// TIA Portal project "1905391_001_000" (V16)

(* hardware
DEVICE "S7-1200 station_1"  S7-1200 Station
   slot 0: "Rack_0"  S7-1200 Rack  Rack  V1.0
   slot 1: "PLC_1"  CPU 1212C DC/DC/Rly  6ES7 212-1HE40-0XB0  V4.4
DEVICE "HMI_1"  TP900 Comfort
   slot 0: "HMI_1"  TP900 Comfort  6AV2 124-0JC01-0AX0  16.0.0.0
   slot 1: "HMI_RT_1"  TP900 Comfort  6AV2 124-0JC01-0AX0  16.0.0.0
   slot 5: "HMI_1.IE_CP_1"  PROFINET Interface  16.0.0.0
      slot 1: "PROFINET Interface_1"  PROFINET Interface
         slot 1: "Port_1"  Port
         slot 2: "Port_2"  Port
   slot 7: "HMI_1.MPI/DP_CP_1"  MPI/DP Interface  16.0.0.0
*)

// ===== PLC "PLC_1"  CPU 1212C DC/DC/Rly =====

VAR_GLOBAL   // PLC tag table "Default tag table"
   "System_Byte" AT %MB1 : Byte;
   "FirstScan" AT %M1.0 : Bool;
   "DiagStatusUpdate" AT %M1.1 : Bool;
   "AlwaysTRUE" AT %M1.2 : Bool;
   "AlwaysFALSE" AT %M1.3 : Bool;
   "Clock_Byte" AT %MB0 : Byte;
   "Clock_10Hz" AT %M0.0 : Bool;
   "Clock_5Hz" AT %M0.1 : Bool;
   "Clock_2.5Hz" AT %M0.2 : Bool;
   "Clock_2Hz" AT %M0.3 : Bool;
   "Clock_1.25Hz" AT %M0.4 : Bool;
   "Clock_1Hz" AT %M0.5 : Bool;
   "Clock_0.625Hz" AT %M0.6 : Bool;
   "Clock_0.5Hz" AT %M0.7 : Bool;
END_VAR

VAR_GLOBAL CONSTANT   // PLC tag table "Default tag table"
   "STRING_LENGTH" : Int := 20;
   "ADP_PARAMETER_LENGTH" : Int := 5;
   "NULL_TOKEN" : Int := -1;
   "BUSY_INDICATOR_OFF" : String := '200;200;200';
   "BUSY_INDICATOR_ON" : String := '250;250;150';
   "ERROR_INDICATOR_OFF" : String := '200;200;200';
   "ERROR_INDICATOR_ON" : String := '250;150;150';
   "STATUS_CODE_OFF" : String := '200;200;200';
   "OPERATION_LABEL_OFF" : String := '200;200;200';
   "CONNECTION_STATUS_HEADER" : String := '200;200;200';
   "STATUS_CODE_PROBLEM" : String := '250;150;150';
   "STATUS_CODE_GOOD" : String := '150;250;150';
END_VAR

VAR_GLOBAL CONSTANT   // PLC tag table "Colors"
   "LABEL_COLOR" : String := '200_200_200';
   "DESELECTED_INPUT_COLOR" : String := '250_250_250';
   "SELECTED_INPUT_COLOR" : String := '150,250,150';
   "BORDER_COLOR" : String := '200_200_200';
   "DIVIDER_COLOR" : String := '50_75_100';
   "THIS_SCREEN_COLOR" : String := '150;150;150';
   "OTHER_SCREEN_COLOR" : String := '100,100,100';
   "ACTUATE" : String := '150_250_150';
   "BACKGROUND_COLOR" : String := '150,150,200';
   "DONE_INDICATOR_OFF" : String := '200;200;200';
   "DONE_INDICATOR_ON" : String := '150;250;150';
   "OPERATION_OFF" : String := '200;200;200';
END_VAR

VAR_GLOBAL CONSTANT   // PLC tag table "Screen_Numbers"
   "WIRE_SCREEN_NUMBER" : Int := 1;
   "MATERIAL_SCREEN_NUMBER" : Int := 2;
   "CONNECTION_CONTROLS_SCREEN_NUMBER" : Int := 3;
   "CONNECTION_STATUS_DETAILS_SCREEN_NUMBER" : Int := 4;
   "CONNECTION_PARAMETERS_SCREEN_NUMBER" : Int := 5;
END_VAR

VAR_GLOBAL CONSTANT   // PLC tag table "Parameter_Entry_Modes"
   "MATERIAL" : String := 'MATERIAL';
   "WIRE" : String := 'WIRE';
END_VAR

VAR_GLOBAL CONSTANT   // PLC tag table "Connection_Statuses"
   "IDLE" : Word := 16#7000;
   "SUCCESS" : Word := 0;
END_VAR

VAR_GLOBAL CONSTANT   // PLC tag table "Send_Modes"
   "MANUAL" : String := 'MANUAL';
   "AUTOMATIC" : String := 'AUTOMATIC';
END_VAR

VAR_GLOBAL CONSTANT   // PLC tag table "Connection_Modes"
   "DISCONNECT_SELECTOR" : DInt := 1;
   "CONNECT_SELECTOR" : DInt := 2;
   "SEND_SELECTOR" : DInt := 3;
   "MATERIAL_DISCONNECT" : DInt := 1;
   "MATERIAL_CONNECT" : DInt := 2;
   "MATERIAL_SEND" : DInt := 3;
   "WIRE_DISCONNECT" : DInt := 4;
   "WIRE_CONNECT" : DInt := 5;
   "WIRE_SEND" : DInt := 6;
END_VAR

TYPE "Divider.UDT"
   STRUCT
      background_animate : DInt;
      background_visible : Bool;
      line_animate : DInt;
      line_visible : Bool;
   END_STRUCT;
END_TYPE

TYPE "Row_Data.UDT"
   STRUCT
      background_animate : DInt;
      background_visible : Bool;
      cell_0_animate : DInt;
      cell_0_visible : Bool;
      cell_1_active : Bool;
      cell_1_animate : DInt;
      cell_1_enable : Bool;
      cell_1_input_finished : Bool;
      cell_1_value : String[50];
      cell_1_visible : Bool;
   END_STRUCT;
END_TYPE

TYPE "HMI_Interface.UDT"
   STRUCT
      connection_parameters : "Connection_Paramters_HMI.UDT";
      connection_status_details : "Connection_Detail.HMI.UDT";
      connection_controls : "Connection_Status.HMI.UDT";
      materials : "Materials.HMI.UDT";
      meta : "HMI_Meta.UDT";
      navigation : "Navigation.HMI.UDT";
      wires : "Wire.HMI.UDT";
   END_STRUCT;
END_TYPE

TYPE "Navigation.HMI.UDT"
   STRUCT
      background_animate : DInt;
      background_visible : Bool;
      bottom_line_animate : DInt;
      bottom_line_visible : Bool;
      communications_status_actuate : Bool;
      communications_status_animate : DInt;
      communications_status_cover_animate : DInt;
      communications_status_cover_visible : Bool;
      communications_status_enable : Bool;
      communications_status_visible : Bool;
      material_actuate : Bool;
      material_animate : DInt;
      material_cover_animate : DInt;
      material_cover_visible : Bool;
      material_enable : Bool;
      material_visible : Bool;
      wire_actuate : Bool;
      wire_animate : DInt;
      wire_cover_animate : DInt;
      wire_cover_visible : Bool;
      wire_enable : Bool;
      wire_visible : Bool;
   END_STRUCT;
END_TYPE

TYPE "Row_Custom.UDT"
   STRUCT
      background_animate : DInt;
      background_visible : Bool;
      cell_0_activate : Bool;
      cell_0_animate : DInt;
      cell_0_enable : Bool;
      cell_0_input_finished : Bool;
      cell_0_value : String[50];
      cell_0_visible : Bool;
      cell_1_activate : Bool;
      cell_1_animate : DInt;
      cell_1_enable : Bool;
      cell_1_input_finished : Bool;
      cell_1_value : String[50];
      cell_1_visible : Bool;
   END_STRUCT;
END_TYPE

TYPE "Row_Label.UDT"
   STRUCT
      background_animate : DInt;
      background_visible : Bool;
      cell_0_animate : DInt;
      cell_0_visible : Bool;
      cell_1_animate : DInt;
      cell_1_visible : Bool;
   END_STRUCT;
END_TYPE

TYPE "HMI_Meta.UDT"
   STRUCT
      screen_number : Int;
      parameter_entry_mode : String;
      connection_mode : DInt;
   END_STRUCT;
END_TYPE

TYPE "Screen_Background.UDT"
   STRUCT
      color : DInt;
      visible : Bool;
   END_STRUCT;
END_TYPE

// folder: LED

TYPE "LED_Interfaces.UDT"
   STRUCT
      material : "LED_Interface.UDT";
      wire : "LED_Interface.UDT";
   END_STRUCT;
END_TYPE

TYPE "LED_Interface.UDT"
   STRUCT
      connection_parameters : "Connection_Parameters.UDT";
      requests : "Connection_Requests.UDT";
      send_buffer : "ADP.Message_Buffer.UDT";
      statuses : "Connection_Statuses.UDT";
   END_STRUCT;
END_TYPE

// folder: adp

TYPE "ADP.Row.2_Cells.UDT"
   STRUCT
      me : Array[0..1] of "ADP.Cell.UDT";
   END_STRUCT;
END_TYPE

TYPE "ADP.Cell.UDT"
   STRUCT
      color : String["ADP_PARAMETER_LENGTH"];
      flashing : String["ADP_PARAMETER_LENGTH"];
      h_align : String["ADP_PARAMETER_LENGTH"];
      line_control : String["ADP_PARAMETER_LENGTH"];
      scroll_speed : String["ADP_PARAMETER_LENGTH"];
      size_and_face : String["ADP_PARAMETER_LENGTH"];
      v_align : String["ADP_PARAMETER_LENGTH"];
      value : String["STRING_LENGTH"];
   END_STRUCT;
END_TYPE

TYPE "ADP.Message_Buffer.UDT"
   STRUCT
      me : Array[0..999] of Byte;
   END_STRUCT;
END_TYPE

TYPE "ADP.Decoded.UDT"
   STRUCT
      color : "ADP.Decoded.Color.UDT";
      flash : "ADP.Decoded.Flash.UDT";
      horizontal_alignment : "ADP.Decoded.Horizontal_Alignment.UDT";
      line_control : "ADP.Decoded.Line_Control.UDT";
      scroll_speed : "ADP.Decoded.Scroll_Speed.UDT";
      size_and_face : "ADP.Decoded.Size_and_Face.UDT";
      vertical_alignment : "ADP.Decoded.Vertical_Alignment.UDT";
   END_STRUCT;
END_TYPE

TYPE "ADP.Decoded.Color.UDT"
   STRUCT
      black : String[8] := 'black';
      blue : String[8] := 'blue';
      green : String[8] := 'green';
      mix_1 : String[8] := 'mix 1';
      mix_2 : String[8] := 'mix 2';
      mix_3 : String[8] := 'mix 3';
      mix_4 : String[8] := 'mix 4';
      red : String[8] := 'red';
      white : String[8] := 'white';
      yellow : String[8] := 'yellow';
   END_STRUCT;
END_TYPE

TYPE "ADP.Decoded.Flash.UDT"
   STRUCT
      off : String[8] := 'off';
      on : String[8] := 'on';
   END_STRUCT;
END_TYPE

TYPE "ADP.Decoded.Horizontal_Alignment.UDT"
   STRUCT
      center : String[8] := 'center';
      left : String[8] := 'left';
      right : String[8] := 'right';
   END_STRUCT;
END_TYPE

TYPE "ADP.Encoded.UDT"
VERSION : 0.1
   STRUCT
      file_system : "ADP.Encoded.File_System.UDT";
      formatting : "ADP.Encoded.Formatting.UDT";
   END_STRUCT;
END_TYPE

TYPE "ADP.Message_Formats.Encoded.UDT"
   STRUCT
      color : String [5];
      flash : String [5];
      scroll_speed : String [5];
      size_and_face : String [5];
      vertical_alignment : String [5];
      horizontal_alignment : String [5];
   END_STRUCT;
END_TYPE

TYPE "ADP.Message_Formats.Decoded.UDT"
   STRUCT
      color : String [20];
      flash : String [20];
      scroll_speed : String [20];
      size_and_face : String [20];
      vertical_alignment : String [20];
      horizontal_alignment : String [20];
   END_STRUCT;
END_TYPE

TYPE "ADP.Decoded.Scroll_Speed.UDT"
   STRUCT
      slowest : String[9] := 'slowest';
      slow : String[9] := 'slow';
      normal : String[9] := 'normal';
      fast : String[9] := 'fast';
      fastest : String[9] := 'fastest';
   END_STRUCT;
END_TYPE

TYPE "ADP.Decoded.Size_and_Face.UDT"
   STRUCT
      bold_5 : String[11] := 'bold 5';
      bold_11 : String[11] := 'bold 11';
      bold_14 : String[11] := 'bold 14';
      bold_15 : String[11] := 'bold 15';
      bold_16 : String[11] := 'bold 16';
      bold_22 : String[11] := 'bold 22';
      bold_30 : String[11] := 'bold 30';
      bold_32 : String[11] := 'bold 32';
      bold_40 : String[11] := 'bold 40';
      normal_5 : String[11] := 'normal 5';
      normal_7 : String[11] := 'normal 7';
      normal_9 : String[11] := 'normal 9';
      normal_11 : String[11] := 'normal 11';
      normal_14 : String[11] := 'normal 14';
      normal_15 : String[11] := 'normal 15';
      normal_16 : String[11] := 'normal 16';
      normal_22 : String[11] := 'normal 22';
      normal_24 : String[11] := 'normal 24';
      normal_30 : String[11] := 'normal 30';
      normal_32 : String[11] := 'normal 32';
      normal_40 : String[11] := 'normal 40';
   END_STRUCT;
END_TYPE

TYPE "ADP.Decoded.Vertical_Alignment.UDT"
   STRUCT
      bottom_hold : String[15] := 'bottom hold';
      fill_hold : String[15] := 'fill hold';
      middle_hold : String[15] := 'middle hold';
      top_hold : String[15] := 'top hold';
      bottom_scroll : String[15] := 'bottom scroll';
      fill_scroll : String[15] := 'fill scroll';
      middle_scroll : String[15] := 'middle scroll';
      top_scroll : String[15] := 'top scroll';
   END_STRUCT;
END_TYPE

TYPE "ADP.Encoded.File_System.UDT"
   STRUCT
      "00 Start of Header" : String[5] := '$01';
      "01 Address" : String[5] := 'Z00';
      "02 Start of Text" : String[5] := '$02';
      "03 Command & File" : String[5] := 'AA';
      "04 END" : String[5] := '$04';
   END_STRUCT;
END_TYPE

TYPE "ADP.Encoded.Formatting.UDT"
   STRUCT
      color : "ADP.Encoded.Formatting.Color.UDT";
      flashing : "ADP.Encoded.Formatting.Flashing.UDT";
      horizontal_alignment : "ADP.Encoded.Formatting.Horizonta_Alignment.UDT";
      line_control : "ADP.Encoded.Formatting.Line_Control.UDT";
      scroll_speed : "ADP.Encoded.Formatting.Scroll_Speed.UDT";
      size_and_face : "ADP.Encoded.Formatting.Size_and_Face.UDT";
      vertical_alignment : "ADP.Encoded.Formatting.Vertical_Alignment.UDT";
   END_STRUCT;
END_TYPE

TYPE "ADP.Encoded.Formatting.Color.UDT"
   STRUCT
      black : String[5] := '$1C0';
      blue : String[5] := '$1C8';
      green : String[5] := '$1C2';
      mix_1 : String[5] := '$1C4';
      mix_2 : String[5] := '$1C5';
      mix_3 : String[5] := '$1C6';
      mix_4 : String[5] := '$1CY';
      red : String[5] := '$1C1';
      white : String[5] := '$1C9';
      yellow : String[5] := '$1C3';
   END_STRUCT;
END_TYPE

TYPE "ADP.Encoded.Formatting.Flashing.UDT"
   STRUCT
      off : String[5] := '$070';
      on : String[5] := '$071';
   END_STRUCT;
END_TYPE

TYPE "ADP.Encoded.Formatting.Size_and_Face.UDT"
   STRUCT
      bold_5 : String[5] := '$1AG';
      bold_11 : String[5] := '$1AH';
      bold_14 : String[5] := '$1A5';
      bold_15 : String[5] := '$1A6';
      bold_16 : String[5] := '$1A7';
      bold_22 : String[5] := '$1AC';
      bold_30 : String[5] := '$1AI';
      bold_32 : String[5] := '$1AJ';
      bold_40 : String[5] := '$1AK';
      normal_5 : String[5] := '$1A0';
      normal_7 : String[5] := '$1A1';
      normal_9 : String[5] := '$1A8';
      normal_11 : String[5] := '$1A9';
      normal_14 : String[5] := '$1A2';
      normal_15 : String[5] := '$1A3';
      normal_16 : String[5] := '$1A4';
      normal_22 : String[5] := '$1AA';
      normal_24 : String[5] := '$1AB';
      normal_30 : String[5] := '$1AD';
      normal_32 : String[5] := '$1AE';
      normal_40 : String[5] := '$1AF';
   END_STRUCT;
END_TYPE

TYPE "ADP.Encoded.Formatting.Horizonta_Alignment.UDT"
   STRUCT
      center : String[5] := '$L1';
      left : String[5] := '$L0';
      right : String[5] := '$L2';
   END_STRUCT;
END_TYPE

TYPE "ADP.Encoded.Formatting.Vertical_Alignment.UDT"
   STRUCT
      middle_hold : String[5] := '$1B b';
      fill_hold : String[5] := '$1B"b';
      bottom_hold : String[5] := '$1B&b';
      top_hold : String[5] := '$1B0b';
      bottom_scroll : String[5] := '$1B a';
      fill_scroll : String[5] := '$1B"a';
      middle_scroll : String[5] := '$1B&a';
      top_scroll : String[5] := '$1B0a';
   END_STRUCT;
END_TYPE

TYPE "ADP.Encoded.Formatting.Scroll_Speed.UDT"
   STRUCT
      slowest : String[5] := '$15';
      slow : String[5] := '$16';
      normal : String[5] := '$17';
      fast : String[5] := '$18';
      fastest : String[5] := '$19';
   END_STRUCT;
END_TYPE

TYPE "ADP.Encoded.Formatting.Line_Control.UDT"
   STRUCT
      new_line : String[5] := '$R';
      word_wrap : String[5] := '';
   END_STRUCT;
END_TYPE

TYPE "ADP.Decoded.Line_Control.UDT"
   STRUCT
      new_line : String[9] := 'new line';
      word_wrap : String[9] := 'word wrap';
   END_STRUCT;
END_TYPE

// folder: connection

TYPE "Connection_Detail.HMI.UDT"
   STRUCT
      back_button_actuate : Bool;
      back_button_enable : Bool;
      back_button_visible : Bool;
      detailed_status_animate : DInt;
      detailed_status_visible : Bool;
      detailed_status_list_selector : DInt;
      detailed_status_message_selector : DInt;
      display_payload_button_actuate : Bool;
      display_payload_button_animate : DInt;
      display_payload_button_enable : Bool;
      display_payload_button_visible : Bool;
      header_animate : DInt;
      header_selector : DInt;
      header_visible : Bool;
      payload_animate : DInt;
      payload_text : String;
      payload_visible : Bool;
   END_STRUCT;
END_TYPE

TYPE "Connection_Requests.UDT"
   STRUCT
      connect : Bool;
      diagnostics : Bool;
      disconnect : Bool;
      reset : Bool;
      send : Bool;
   END_STRUCT;
END_TYPE

TYPE "Connection_Parameters.UDT"
   STRUCT
      id : Conn_Ouc;
      ip_address : String[15];
      port_number : String[15];
   END_STRUCT;
END_TYPE

TYPE "Connection_Parameters_HMI_Interface.UDT"
   STRUCT
      back_actuate : Bool;
      back_animate : DInt;
      back_enable : Bool;
      back_visible : Bool;
      header_animate : DInt;
      header_value : String[25];
      header_visible : Bool;
      id_label_animate : DInt;
      id_label_visible : Bool;
      id_entry_active : Bool;
      id_entry_animate : DInt;
      id_entry_input_finished : Bool;
      id_entry_enable : Bool;
      id_entry_value : String[6];
      id_entry_visible : Bool;
      ip_address_label_animate : DInt;
      ip_address_label_visible : Bool;
      ip_address_entry_active : Bool;
      ip_address_entry_animate : DInt;
      ip_address_entry_enable : Bool;
      ip_address_entry_input_finished : Bool;
      ip_address_entry_value : String[15];
      ip_address_entry_visible : Bool;
      port_label_animate : DInt;
      port_label_visible : Bool;
      port_entry_active : Bool;
      port_entry_animate : DInt;
      port_entry_enable : Bool;
      port_entry_input_finished : Bool;
      port_entry_value : String[6];
      port_entry_visible : Bool;
   END_STRUCT;
END_TYPE

TYPE "Connection_Paramters_HMI.UDT"
   STRUCT
      background : "Screen_Background.UDT";
      connection_parameters : "Connection_Parameters_HMI_Interface.UDT";
   END_STRUCT;
END_TYPE

// folder: connection/connection_status

TYPE "Connection_Status_Header.UDT"
   STRUCT
      actuate : Bool;
      animate : DInt;
      enable : Bool;
      visible : Bool;
   END_STRUCT;
END_TYPE

TYPE "Connection_Status_Element.UDT"
   STRUCT
      busy_status_indicator_animate : DInt;
      busy_status_indicator_visible : Bool;
      done_status_indicator_animate : DInt;
      done_status_indicator_visible : Bool;
      error_status_indicator_animate : DInt;
      error_status_indicator_visible : Bool;
      operation_button_actuate : Bool;
      operation_button_enable : Bool;
      operation_button_visible : Bool;
      operation_label_animate : DInt;
      operation_label_visible : Bool;
      show_status_code_description_button_actuate : Bool;
      show_status_code_description_button_enable : Bool;
      show_status_code_description_button_visible : Bool;
      status_code_description_animate : DInt;
      status_code_description_value : DInt := -1;
      status_code_description_visible : Bool;
      status_code_label_animate : DInt;
      status_code_label_visible : Bool;
      status_code_value_animate : DInt;
      status_code_value_visible : Bool;
      status_code_value : String[6];
   END_STRUCT;
END_TYPE

TYPE "Connection_Status_Table.UDT"
   STRUCT
      header : "Connection_Status_Header.UDT";
      disconnect : "Connection_Status_Element.UDT";
      connect : "Connection_Status_Element.UDT";
      send : "Connection_Status_Element.UDT";
   END_STRUCT;
END_TYPE

TYPE "Connection_Status.HMI.UDT"
   STRUCT
      background : "Screen_Background.UDT";
      material : "Connection_Status_Table.UDT";
      wire : "Connection_Status_Table.UDT";
   END_STRUCT;
END_TYPE

TYPE "Connection_Status.UDT"
   STRUCT
      done : Bool;
      busy : Bool;
      error : Bool;
      status : Word;
   END_STRUCT;
END_TYPE

TYPE "Connection_Statuses.UDT"
   STRUCT
      diagnostics : "Connection_Status.UDT";
      disconnect : "Connection_Status.UDT";
      connect : "Connection_Status.UDT";
      reset : "Connection_Status.UDT";
      send : "Connection_Status.UDT";
   END_STRUCT;
END_TYPE

TYPE "Connection_Status_Timers.UDT"
   STRUCT
      busy : TOF_TIME;
      error : TOF_TIME;
      status : TOF_TIME;
   END_STRUCT;
END_TYPE

// folder: material

TYPE "Materials.HMI.UDT"
   STRUCT
      background : "Screen_Background.UDT";
      bottom_border : "Divider.UDT";
      chromium : "Row_Data.UDT";
      custom : "Row_Custom.UDT";
      divider : "Divider.UDT";
      header : "Row_Label.UDT";
      heat : "Row_Data.UDT";
      manganese : "Row_Data.UDT";
      molybdenum : "Row_Data.UDT";
      nickel : "Row_Data.UDT";
      silicon : "Row_Data.UDT";
      vanadium : "Row_Data.UDT";
   END_STRUCT;
END_TYPE

TYPE "Material.Data.UDT"
   STRUCT
      chromium : Real;
      custom_value : Real;
      custom_name : String[50];
      heat : Real;
      manganese : Real;
      molybdenum : Real;
      nickel : Real;
      silicon : Real;
      vanadium : Real;
   END_STRUCT;
END_TYPE

// folder: wire

TYPE "Wire.UDT"
   STRUCT
      aluminum : Real;
      calcium_silicon : Real;
      carbon : Real;
      custom : Real;
      heat : Real;
      sulfur : Real;
   END_STRUCT;
END_TYPE

TYPE "Wire.HMI.UDT"
   STRUCT
      aluminum : "Row_Data.UDT";
      background : "Screen_Background.UDT";
      bottom_border : "Divider.UDT";
      calcium_silicon : "Row_Data.UDT";
      carbon : "Row_Data.UDT";
      divider : "Divider.UDT";
      header : "Row_Label.UDT";
      heat : "Row_Data.UDT";
      sulfur : "Row_Data.UDT";
   END_STRUCT;
END_TYPE

// folder: 00/data

DATA_BLOCK "ADP_Library"   // DB1
{ S7_Optimized_Access := 'TRUE' }
VERSION : 0.1
BEGIN
END_DATA_BLOCK

DATA_BLOCK "HMI_Interface.Data"   // DB2
{ S7_Optimized_Access := 'TRUE' }
VERSION : 0.1
BEGIN
   meta.screen_number := 1;
END_DATA_BLOCK

DATA_BLOCK "LED_Interface.Data"   // DB3
{ S7_Optimized_Access := 'TRUE' }
VERSION : 0.1
BEGIN
END_DATA_BLOCK

DATA_BLOCK "Display_IDB"   // DB4
{ S7_Optimized_Access := 'TRUE' }
VERSION : 0.1
// stored: InstanceOfName Display
"Display"
BEGIN
END_DATA_BLOCK

DATA_BLOCK "Middleware_IDB"   // DB5
{ S7_Optimized_Access := 'TRUE' }
VERSION : 0.1
// stored: InstanceOfName Middleware
"Middleware"
BEGIN
END_DATA_BLOCK

// folder: (top level)

ORGANIZATION_BLOCK "Main"   // OB1, LAD, ProgramCycle
TITLE = "Main Program Sweep (Cycle)"
{ S7_Optimized_Access := 'TRUE' }
VERSION : 0.1
   VAR_INPUT
      Initial_Call : Bool;   // Initial call of this OB
      Remanence : Bool;   // =True, if remanent data are available
   END_VAR
BEGIN

REGION Network 1
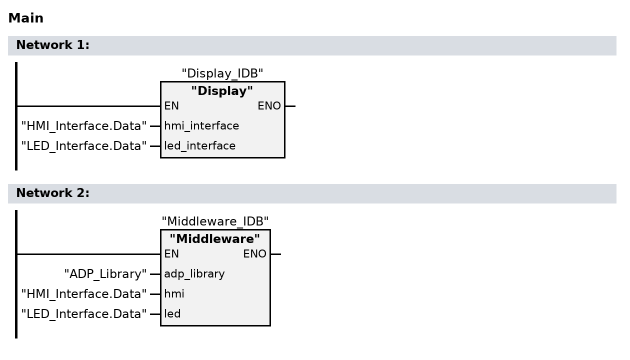
   RUNG wire#powerrail
      "Display_IDB"(hmi_interface := "HMI_Interface.Data", led_interface := "LED_Interface.Data")
   END_RUNG
   // the same network as SCL:
   "Display_IDB"(hmi_interface := "HMI_Interface.Data", led_interface := "LED_Interface.Data");   // "Display"
END_REGION

REGION Network 2
   RUNG wire#powerrail
      "Middleware_IDB"(adp_library := "ADP_Library", hmi := "HMI_Interface.Data", led := "LED_Interface.Data")
   END_RUNG
   // the same network as SCL:
   "Middleware_IDB"(adp_library := "ADP_Library", hmi := "HMI_Interface.Data", led := "LED_Interface.Data");   // "Middleware"
END_REGION
END_ORGANIZATION_BLOCK

ORGANIZATION_BLOCK "Time error interrupt"   // OB80, LAD, TimeErrorInterrupt
{ S7_Optimized_Access := 'TRUE' }
VERSION : 0.1
   VAR_INPUT
      Fault_ID : Byte;   // Fault identifier
      Csg_OBnr : OB_Any;   // Number of OB causing the error
      Csg_Prio : UInt;   // Priority of OB causing the error
   END_VAR
BEGIN
END_ORGANIZATION_BLOCK

ORGANIZATION_BLOCK "Startup"   // OB100, LAD, Startup
TITLE = "Complete Restart"
{ S7_Optimized_Access := 'TRUE' }
VERSION : 0.1
   VAR_INPUT
      LostRetentive : Bool;   // True if retentive data are lost
      LostRTC : Bool;   // True if date and time are lost
   END_VAR
BEGIN

REGION Network 1: INITIALIZE MATERIALS PAGE
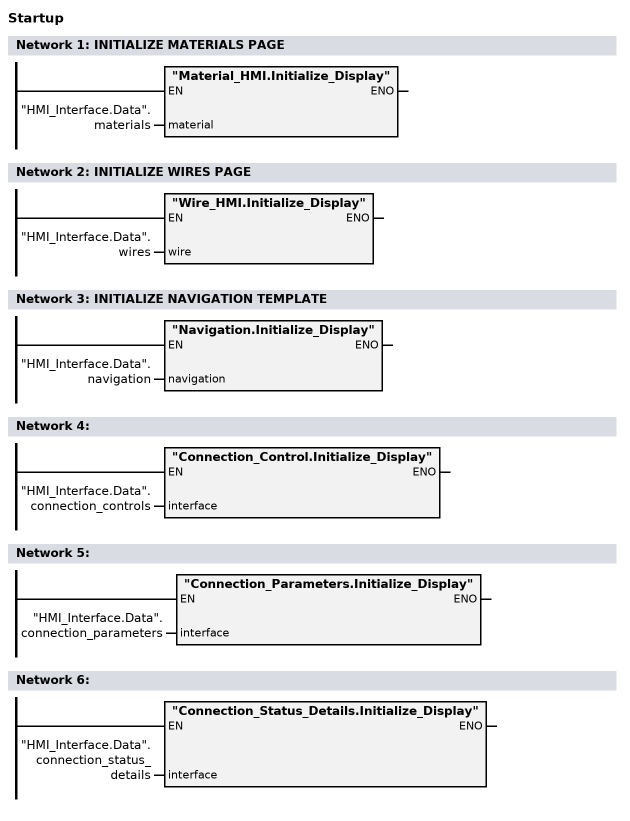
   RUNG wire#powerrail
      "Material_HMI.Initialize_Display"(material := "HMI_Interface.Data".materials)
   END_RUNG
   // the same network as SCL:
   "Material_HMI.Initialize_Display"(material := "HMI_Interface.Data".materials);
END_REGION

REGION Network 2: INITIALIZE WIRES PAGE
   RUNG wire#powerrail
      "Wire_HMI.Initialize_Display"(wire := "HMI_Interface.Data".wires)
   END_RUNG
   // the same network as SCL:
   "Wire_HMI.Initialize_Display"(wire := "HMI_Interface.Data".wires);
END_REGION

REGION Network 3: INITIALIZE NAVIGATION TEMPLATE
   RUNG wire#powerrail
      "Navigation.Initialize_Display"(navigation := "HMI_Interface.Data".navigation)
   END_RUNG
   // the same network as SCL:
   "Navigation.Initialize_Display"(navigation := "HMI_Interface.Data".navigation);
END_REGION

REGION Network 4
   RUNG wire#powerrail
      "Connection_Control.Initialize_Display"(interface := "HMI_Interface.Data".connection_controls)
   END_RUNG
   // the same network as SCL:
   "Connection_Control.Initialize_Display"(interface := "HMI_Interface.Data".connection_controls);
END_REGION

REGION Network 5
   RUNG wire#powerrail
      "Connection_Parameters.Initialize_Display"(interface := "HMI_Interface.Data".connection_parameters)
   END_RUNG
   // the same network as SCL:
   "Connection_Parameters.Initialize_Display"(interface := "HMI_Interface.Data".connection_parameters);
END_REGION

REGION Network 6
   RUNG wire#powerrail
      "Connection_Status_Details.Initialize_Display"(interface := "HMI_Interface.Data".connection_status_details)
   END_RUNG
   // the same network as SCL:
   "Connection_Status_Details.Initialize_Display"(interface := "HMI_Interface.Data".connection_status_details);
END_REGION
END_ORGANIZATION_BLOCK

// folder: 00/display

FUNCTION_BLOCK "Display"   // FB5, SCL
{ S7_Optimized_Access := 'TRUE' }
VERSION : 0.1
   VAR_IN_OUT
      hmi_interface : "HMI_Interface.UDT";
      led_interface : "LED_Interfaces.UDT";
   END_VAR
   VAR
      hmi_display : "HMI";
      material_led : "Sign.Connection";
      wire_led : "Sign.Connection";
   END_VAR
BEGIN
   REGION "HMI"
       #hmi_display(led_interface := #led_interface,
                    hmi_interface := #hmi_interface);
   END_REGION


   REGION "LED"
       #material_led(#led_interface.material);
       #wire_led(#led_interface.wire);
   END_REGION
END_FUNCTION_BLOCK

// folder: 00/middleware

FUNCTION_BLOCK "Middleware"   // FB2, SCL
{ S7_Optimized_Access := 'TRUE' }
VERSION : 0.1
   VAR_INPUT
      adp_library : "ADP.Encoded.UDT";
   END_VAR
   VAR_IN_OUT
      hmi : "HMI_Interface.UDT";
      led : "LED_Interfaces.UDT";
   END_VAR
   VAR
      material_messaging : "Material_Message";
      wire_messaging : "Wire_Message";
   END_VAR
BEGIN
   REGION "PROCESS CONNECTION PARAMETER INPUTS"
       IF #hmi.meta.screen_number = "CONNECTION_PARAMETERS_SCREEN_NUMBER" THEN
           "Material_Sign.Set_Connection_Parameters"(mode := #hmi.meta.parameter_entry_mode,
                                                     interface := #hmi.connection_parameters.connection_parameters,
                                                     saved := #led.material.connection_parameters);
           "Wire_Sign.Set_Connection_Parameters"(mode := #hmi.meta.parameter_entry_mode,
                                                 interface := #hmi.connection_parameters.connection_parameters,
                                                 saved := #led.wire.connection_parameters);
       END_IF;
   END_REGION


   REGION "MESSAGE DRIVER FOR MATERIALS SIGN"
       #material_messaging(adp_liberary := #adp_library,
                           hmi_interface := #hmi,
                           led_interface := #led.material);
   END_REGION

   REGION "WIRE MESSAGE ASSEMBLY AND SEND REQUESTS ORIGINATION"
       #wire_messaging(adp_liberary := #adp_library,
                       hmi_interface := #hmi,
                       led_interface := #led.wire);
   END_REGION
END_FUNCTION_BLOCK

// folder: HMI

FUNCTION_BLOCK "HMI"   // FB6, SCL
{ S7_Optimized_Access := 'TRUE' }
VERSION : 0.1
   VAR_IN_OUT
      hmi_interface : "HMI_Interface.UDT";
      led_interface : "LED_Interfaces.UDT";
   END_VAR
   VAR
      material_requests : "Connection.Requests";
      wire_requests : "Connection.Requests";
   END_VAR
BEGIN
   "HMI.Navigation_Screen"(interface := #hmi_interface);

   CASE #hmi_interface.meta.screen_number OF

       "MATERIAL_SCREEN_NUMBER":
           "HMI.Material_Screen"(#hmi_interface.materials);

       "WIRE_SCREEN_NUMBER":
           "HMI.Wire_Screen"(#hmi_interface.wires);

       "CONNECTION_CONTROLS_SCREEN_NUMBER":
           "HMI.Connection_Controls_Screen"(led_interface := #led_interface,
                                            hmi_interface := #hmi_interface,
                                            material_requests := #material_requests,
                                            wire_requests := #wire_requests);

       "CONNECTION_PARAMETERS_SCREEN_NUMBER":
           "HMI.Connection_Parameters_Screen"(hmi_interface := #hmi_interface,
                                              led_interface := #led_interface,
                                              interface := #hmi_interface.connection_parameters);

       "CONNECTION_STATUS_DETAILS_SCREEN_NUMBER":
           "HMI.Connection_Status_Details_Screen"(led_interfaces := #led_interface,
                                                  meta := #hmi_interface.meta,
                                                  interface := #hmi_interface.connection_status_details);

   END_CASE;
END_FUNCTION_BLOCK

FUNCTION "HMI.Wire_Screen" : Void   // FC3, SCL
{ S7_Optimized_Access := 'TRUE' }
VERSION : 0.1
   VAR_IN_OUT
      wire : "Wire.HMI.UDT";
   END_VAR
BEGIN
   "Wire_HMI.Input_Animations"(#wire);
END_FUNCTION

FUNCTION "HMI.Material_Screen" : Void   // FC4, SCL
{ S7_Optimized_Access := 'TRUE' }
VERSION : 0.1
   VAR_IN_OUT
      material : "Materials.HMI.UDT";
   END_VAR
BEGIN
   "Material_HMI.Input_Animations"(#material);
END_FUNCTION

FUNCTION "HMI.Navigation_Screen" : Void   // FC8, SCL
{ S7_Optimized_Access := 'TRUE' }
VERSION : 0.1
   VAR_IN_OUT
      interface : "HMI_Interface.UDT";
   END_VAR
BEGIN
   "Navigation.Material_Animation"(screen_number := #interface.meta.screen_number,
                                             navigation := #interface.navigation);
   "Navigation.Wire_Animation"(screen_number := #interface.meta.screen_number,
                                         navigation := #interface.navigation);
   "Navigation.Bottom_Cover_Animations"(screen_number := #interface.meta.screen_number,
                                        navigation := #interface.navigation);
   "Navigation.Connections_Screen_Animation"(screen_number := #interface.meta.screen_number,
                                                          navigation := #interface.navigation);
END_FUNCTION

FUNCTION "HMI.Connection_Controls_Screen" : Void   // FC84, SCL
{ S7_Optimized_Access := 'TRUE' }
VERSION : 0.1
   VAR_IN_OUT
      hmi_interface : "HMI_Interface.UDT";
      led_interface : "LED_Interfaces.UDT";
      material_requests : "Connection.Requests";
      wire_requests : "Connection.Requests";
   END_VAR
BEGIN
   REGION "ANIMATIONS"
       "Connection_Control_Table.Animate"(statuses := #led_interface.material.statuses,
                                          interface := #hmi_interface.connection_controls.material);
       "Connection_Control_Table.Animate"(statuses := #led_interface.wire.statuses,
                                          interface := #hmi_interface.connection_controls.wire);
   END_REGION


   REGION "SET GLOBAL MODES"
       "Connection_Parameters.Set_Mode"(interface := #hmi_interface.connection_controls,
                                        meta := #hmi_interface.meta);
       "Connection_Status_Details.Set_Mode"(interface := #hmi_interface.connection_controls,
                                            mode := #hmi_interface.meta.connection_mode);
   END_REGION


   REGION "CONNECTION REQUESTS"
       #material_requests(hmi := #hmi_interface.connection_controls.material,
                          sign := #led_interface.material.requests);
       #wire_requests(hmi := #hmi_interface.connection_controls.wire,
                      sign := #led_interface.wire.requests);
   END_REGION


   REGION "LOAD CONNECTION PARAMETER INFORMATION"
       IF #hmi_interface.connection_controls.material.header.actuate OR #hmi_interface.connection_controls.wire.header.actuate THEN
           "Connection_Parameters.Reload_Screen"(meta := #hmi_interface.meta,
                                                 connection_controls := #hmi_interface.connection_controls,
                                                 led := #led_interface,
                                                 hmi := #hmi_interface.connection_parameters);
       END_IF;
   END_REGION
END_FUNCTION

FUNCTION "HMI.Connection_Parameters_Screen" : Void   // FC131, SCL
{ S7_Optimized_Access := 'TRUE' }
VERSION : 0.1
   VAR_INPUT
      hmi_interface : "HMI_Interface.UDT";
      led_interface : "LED_Interfaces.UDT";
   END_VAR
   VAR_IN_OUT
      interface : "Connection_Paramters_HMI.UDT";
   END_VAR
BEGIN
   REGION "ANIMATIONS"
       "Connection_Parameters.Animate_Back"(#interface.connection_parameters);
       "Connection_Parameters.Animate_ID_Active"(#interface.connection_parameters);
       "Connection_Parameters.Animate_IP_Active"(#interface.connection_parameters);
       "Connection_Parameters.Animate_Port_Active"(#interface.connection_parameters);
   END_REGION
END_FUNCTION

FUNCTION "HMI.Connection_Status_Details_Screen" : Void   // FC164, SCL
{ S7_Optimized_Access := 'TRUE' }
VERSION : 0.1
   VAR_INPUT
      led_interfaces : "LED_Interfaces.UDT";
      meta : "HMI_Meta.UDT";
   END_VAR
   VAR_IN_OUT
      interface : "Connection_Detail.HMI.UDT";
   END_VAR
BEGIN
   "Connection_Status_Details.Set_Header_Selector"(meta := #meta,
                                                   interface := #interface);
   "Connection_Status_Details.Set_Status_Details_Selector"(led_interfaces := #led_interfaces,
                                                           hmi_meta := #meta,
                                                           interface := #interface);

   IF #interface.display_payload_button_actuate THEN
       "Connection_Status_Details.Show_Payload"(led_interfaces := #led_interfaces,
                                                hmi_meta := #meta,
                                                interface := #interface);
       RETURN;
   END_IF;

   "Connection_Status_Details.Display_Detailed_Status"(#interface);
END_FUNCTION

// folder: adp

FUNCTION "ADP.Buffer_to_String" : String   // FC192, SCL
{ S7_Optimized_Access := 'TRUE' }
VERSION : 0.1
   VAR_INPUT
      buffer : "ADP.Message_Buffer.UDT";
      lenWrap : Int;
   END_VAR
   VAR_TEMP
      outBox : String;
      pSerialize : DInt;
      statSerialize : Int;
      byteBox : Array[0..#uBound] of Byte;
      i : Int;
      pByteBox : Int;
      validChar : Bool;
      ofstLabel : DInt;
      stringBox : String;
      remainder : Int;
   END_VAR
   VAR CONSTANT
      all : USInt := 0;
      hex01 : String := '<0x01>';
      hex02 : String := '<0x02>';
      hex04 : String := '<0x04>';
      hex15 : String := '<0x015>';
      hex16 : String := '<0x016>';
      hex17 : String := '<0x017>';
      hex18 : String := '<0x018>';
      hex19 : String := '<0x019>';
      hex1A : String := '<0x1A>';
      hex1B : String := '<0x1B>';
      hex1C : String := '<0x1C>';
      uBound : Int := 999;
      lenLabel : Int := 6;
      lineBreak : Byte := '$L';
   END_VAR
BEGIN
   REGION "SCRUB ARRAY"    
       FOR #i := 0 TO 999 DO

           IF #i > #lenWrap THEN
               Chars_TO_Strg(Chars := #byteBox,
                             pChars := 0,
                             Cnt := #all,
                             Strg => #"ADP.Buffer_to_String");
               RETURN;
           END_IF;

           #validChar := TRUE;

           IF #buffer.me[#i] = 16#01 THEN
               #stringBox := #hex01;
               #validChar := FALSE;
           END_IF;

           IF #buffer.me[#i] = 16#02 THEN
               #stringBox := #hex02;
               #validChar := FALSE;
           END_IF;

           IF #buffer.me[#i] = 16#04 THEN
               #stringBox := #hex04;
               #validChar := FALSE;
           END_IF;

           IF #buffer.me[#i] = 16#15 THEN
               #stringBox := #hex15;
               #validChar := FALSE;
           END_IF;

           IF #buffer.me[#i] = 16#16 THEN
               #stringBox := #hex16;
               #validChar := FALSE;
           END_IF;

           IF #buffer.me[#i] = 16#17 THEN
               #stringBox := #hex17;
               #validChar := FALSE;
           END_IF;

           IF #buffer.me[#i] = 16#18 THEN
               #stringBox := #hex18;
               #validChar := FALSE;
           END_IF;

           IF #buffer.me[#i] = 16#19 THEN
               #stringBox := #hex19;
               #validChar := FALSE;
           END_IF;

           IF #buffer.me[#i] = 16#1A THEN
               #stringBox := #hex1A;
               #validChar := FALSE;
           END_IF;

           IF #buffer.me[#i] = 16#1B THEN
               #stringBox := #hex1B;
               #validChar := FALSE;
           END_IF;

           IF #buffer.me[#i] = 16#1C THEN
               #stringBox := #hex1C;
               #validChar := FALSE;
           END_IF;

           IF NOT #validChar THEN
               #remainder := #pByteBox MOD #lenWrap;
               IF #remainder + #lenLabel > #lenWrap THEN
                   #byteBox[#pByteBox] := #lineBreak;
                   #pByteBox += 1;
               END_IF;
               Strg_TO_Chars(Strg := #stringBox,
                             pChars := #pByteBox,
                             Cnt => #ofstLabel,
                             Chars := #byteBox);
               #pByteBox += DINT_TO_INT(#ofstLabel);
           END_IF;

           IF #validChar THEN
               #byteBox[#pByteBox] := #buffer.me[#i];
               #pByteBox += 1;
           END_IF;

       END_FOR;
   END_REGION

   REGION "CONVERT SCRUBBED ARRAY TO STRING"
       Chars_TO_Strg(Chars := #byteBox,
                     pChars := 0,
                     Cnt := #all,
                     Strg => #"ADP.Buffer_to_String");
   END_REGION
END_FUNCTION

// folder: any_data_types

FUNCTION "Any.Array.Length" : UDInt   // FC16, SCL
{ S7_Optimized_Access := 'TRUE' }
VERSION : 0.1
   VAR_INPUT
      "array" : Variant;
   END_VAR
   VAR_TEMP
      status : DInt;
      ret : UDInt;
   END_VAR
BEGIN
   #ret := CountOfElements(#array);
   #"Any.Array.Length" := #ret;
END_FUNCTION

// folder: bool

FUNCTION "Bool.Animate" : Void   // FC49, SCL
{ S7_Optimized_Access := 'TRUE' }
VERSION : 0.1
   VAR_INPUT
      signal : Bool;
      color_on : DInt;
      color_off : DInt;
   END_VAR
   VAR_IN_OUT
      animation : DInt;
   END_VAR
BEGIN
   IF #signal THEN
       #animation := #color_on;
       RETURN;
   END_IF;
   #animation := #color_off;
   RETURN;
END_FUNCTION

FUNCTION "Bool.Rising_Edge" : Bool   // FC105, SCL
{ S7_Optimized_Access := 'TRUE' }
VERSION : 0.1
   VAR_INPUT
      signal : Bool;
      old_signal : Bool;
   END_VAR
BEGIN
   #"Bool.Rising_Edge" := #signal AND NOT #old_signal;
END_FUNCTION

FUNCTION "Bool.Falling_Edge" : Bool   // FC106, SCL
{ S7_Optimized_Access := 'TRUE' }
VERSION : 0.1
   VAR_INPUT
      signal : Bool;
      old_signal : Bool;
   END_VAR
BEGIN
   #"Bool.Falling_Edge" := NOT #signal AND #old_signal;
END_FUNCTION

// folder: byte

FUNCTION "Byte.to_String" : String   // FC117, SCL
{ S7_Optimized_Access := 'TRUE' }
VERSION : 0.1
   VAR_INPUT
      value : Byte;
   END_VAR
   VAR_TEMP
      _low_nibble : Byte;
      _high_nibble : Byte;
   END_VAR
   VAR CONSTANT
      LOW_NIBBLE_MASK : Byte := 16#0F;
      HIGH_NIBBLE_MASK : Byte := 16#F0;
   END_VAR
BEGIN
   #_low_nibble := #value AND #LOW_NIBBLE_MASK;
   #_high_nibble := SHR_BYTE(IN := #value AND #HIGH_NIBBLE_MASK,
                             N := 4);
   #"Byte.to_String" := CONCAT_STRING(IN1 := "Nibble.to_String"(#_high_nibble),
                                      IN2 := "Nibble.to_String"(#_low_nibble));
END_FUNCTION

// folder: char

FUNCTION "Char.Is_Numeric" : Bool   // FC57, SCL
{ S7_Optimized_Access := 'TRUE' }
VERSION : 0.1
   VAR_INPUT
      character : Char;
   END_VAR
   VAR CONSTANT
      NUMBERS : String := '0123456789';
   END_VAR
BEGIN
   IF FIND(IN1 := #NUMBERS, IN2 := CHAR_TO_STRING(#character)) = 0 THEN
       #"Char.Is_Numeric" := FALSE;
       RETURN;
   END_IF;
   #"Char.Is_Numeric" := TRUE;
   RETURN;
END_FUNCTION

// folder: color

FUNCTION "Color.String_to_DInt" : DInt   // FC14, SCL
{ S7_Optimized_Access := 'TRUE' }
VERSION : 0.1
   VAR_INPUT
      color : String;   // enter rgb value with comma, semicolon, or underscore as delimeter. e.g.: '200,100,200' or '195_168_0'
   END_VAR
   VAR_TEMP
      _color : String;
      _background : DInt;
      _blue : DInt;
      _delimeters : Array[0..2] of String;
      _flash : DInt;
      _green : DInt;
      _red : DInt;
      _substrings : Array[0..3] of String;
   END_VAR
BEGIN
   REGION "COPY TO LOCAL"
       #_color := #color;
   END_REGION


   REGION "BACKGROUND MODE"
       #_background := 1;
       IF "Color.String_Is_Background"(#color) THEN
           #_background := -1;
           #_color := "String.Slice_Right"("string" := #_color,
                                           start_at := 1);
       END_IF;
   END_REGION


   REGION "SET UP DELIMETERS"
       #_delimeters[0] := ',';
       #_delimeters[1] := ';';
       #_delimeters[2] := '_';
   END_REGION


   REGION "SPLIT STRING"
       "String.Split_Multiple"(string_in := #_color,
                               delimeters := #_delimeters,
                               "pointer" := 0,
                               substrings => #_substrings);
       "String.Reverse_Array"(null_token := '',
                              string_array := #_substrings);
   END_REGION


   REGION "RETURN 0 ON INVALID STRING"
       IF NOT "Color.Validate_String"(#_substrings) THEN
           #"Color.String_to_DInt" := 0;
           RETURN;
       END_IF;
   END_REGION


   REGION "CALCULATE CODE"
       #_flash := STRING_TO_DINT(#_substrings[3]) * 1_000_000_000;
       #_red := STRING_TO_DINT(#_substrings[2]) * 1_000_000;
       #_green := STRING_TO_DINT(#_substrings[1]) * 1_000;
       #_blue := STRING_TO_DINT(#_substrings[0]);
   END_REGION


   REGION "RETURN"
       #"Color.String_to_DInt" := #_background * (#_flash + #_red + #_green + #_blue);
       RETURN;
   END_REGION
END_FUNCTION

FUNCTION "Color.Set_As_Background" : DInt   // FC27, SCL
{ S7_Optimized_Access := 'TRUE' }
VERSION : 0.1
   VAR_INPUT
      color_code : DInt;
   END_VAR
BEGIN
   IF #color_code < 0 THEN
       #"Color.Set_As_Background" := -1 * #color_code;
       RETURN;
   END_IF;
   #"Color.Set_As_Background" := #color_code;
   RETURN;
END_FUNCTION

FUNCTION "Color.Set_As_Foreground" : DInt   // FC30, SCL
{ S7_Optimized_Access := 'TRUE' }
VERSION : 0.1
   VAR_INPUT
      color_code : DInt;
   END_VAR
BEGIN
   IF #color_code >= 0 THEN
       #"Color.Set_As_Foreground" := -1 * #color_code;
       RETURN;
   END_IF;
   #"Color.Set_As_Foreground" := #color_code;
   RETURN;
END_FUNCTION

FUNCTION "Color.Flash_On" : DInt   // FC31, SCL
{ S7_Optimized_Access := 'TRUE' }
VERSION : 0.1
   VAR_INPUT
      color_code : DInt;
   END_VAR
   VAR CONSTANT
      FLASH : DInt := 1_000_000_000;
   END_VAR
BEGIN
   #"Color.Flash_On" := #FLASH + #color_code MOD #FLASH;
END_FUNCTION

FUNCTION "Color.Flash_Off" : DInt   // FC32, SCL
{ S7_Optimized_Access := 'TRUE' }
VERSION : 0.1
   VAR_INPUT
      color_code : DInt;
   END_VAR
   VAR CONSTANT
      FLASH : DInt := 1_000_000_000;
   END_VAR
BEGIN
   #"Color.Flash_Off" := #color_code MOD #FLASH;
END_FUNCTION

FUNCTION "Color.String_Is_Background" : Bool   // FC52, SCL
{ S7_Optimized_Access := 'TRUE' }
VERSION : 0.1
   VAR_INPUT
      color : String;
   END_VAR
BEGIN
   IF LEFT(IN := #color, L := 1) = '-' THEN
       #"Color.String_Is_Background" := TRUE;
       RETURN;
   END_IF;
   #"Color.String_Is_Background" := FALSE;
   RETURN;
END_FUNCTION

FUNCTION "Color.DInt_Is_Background" : Bool   // FC53, SCL
{ S7_Optimized_Access := 'TRUE' }
VERSION : 0.1
   VAR_INPUT
      color : DInt;
   END_VAR
BEGIN
   IF #color < 0 THEN
       #"Color.DInt_Is_Background" := FALSE;
       RETURN;
   END_IF;
   #"Color.DInt_Is_Background" := TRUE;
   RETURN;
END_FUNCTION

FUNCTION "Color.DInt_Is_Flashing" : Bool   // FC54, SCL
{ S7_Optimized_Access := 'TRUE' }
VERSION : 0.1
   VAR_INPUT
      color : DInt;
   END_VAR
   VAR CONSTANT
      FLASH : DInt := 1_000_000_000;
   END_VAR
BEGIN
   IF #color / #FLASH > 0 THEN
       #"Color.DInt_Is_Flashing" := TRUE;
       RETURN;
   END_IF;
   #"Color.DInt_Is_Flashing" := FALSE;
   RETURN;
END_FUNCTION

FUNCTION "Color.String_Is_Flashing" : Void   // FC55, SCL
{ S7_Optimized_Access := 'TRUE' }
VERSION : 0.1
   VAR_INPUT
      color : String;
   END_VAR
BEGIN
END_FUNCTION

FUNCTION "Color.Validate_String" : Bool   // FC56, SCL
{ S7_Optimized_Access := 'TRUE' }
VERSION : 0.1
   VAR_INPUT
      color : Array[*] of String;
   END_VAR
   VAR_TEMP
      _i : UDInt;
      _length : UDInt;
   END_VAR
BEGIN
   REGION "INVALID FLASH"
       IF #color[3] <> '1' AND #color[3] <> '' THEN
           #"Color.Validate_String" := FALSE;
           RETURN;
       END_IF;
   END_REGION


   REGION "NON-NUMERIC COMPONENT"
       FOR #_i := 0 TO #_length DO
           IF NOT "String.Is_Numeric"(#color[#_i]) THEN
               #"Color.Validate_String" := FALSE;
               RETURN;
           END_IF;
       END_FOR;
   END_REGION


   REGION "IS VALID"
       #"Color.Validate_String" := TRUE;
       RETURN;
   END_REGION
END_FUNCTION

// folder: divider

FUNCTION "Divider.Show" : Void   // FC2, SCL
{ S7_Optimized_Access := 'TRUE' }
VERSION : 0.1
   VAR_IN_OUT
      divider : "Divider.UDT";
   END_VAR
   VAR CONSTANT
      MODE : Bool := TRUE;
   END_VAR
BEGIN
   #divider.background_visible := #MODE;
   #divider.line_visible := #MODE;
END_FUNCTION

FUNCTION "Divider.Hide_Line" : Void   // FC13, SCL
{ S7_Optimized_Access := 'TRUE' }
VERSION : 0.1
   VAR_IN_OUT
      divider : "Divider.UDT";
   END_VAR
   VAR CONSTANT
      MODE : Bool := FALSE;
   END_VAR
BEGIN
   #divider.line_visible := #MODE;
END_FUNCTION

FUNCTION "Divider.Hide" : Void   // FC19, SCL
{ S7_Optimized_Access := 'TRUE' }
VERSION : 0.1
   VAR_IN_OUT
      divider : "Divider.UDT";
   END_VAR
   VAR CONSTANT
      MODE : Bool := FALSE;
   END_VAR
BEGIN
   #divider.background_visible := #MODE;
   #divider.line_visible := #MODE;
END_FUNCTION

FUNCTION "Divider.Initialize_Colors" : Void   // FC45, SCL
{ S7_Optimized_Access := 'TRUE' }
VERSION : 0.1
   VAR_IN_OUT
      divider : "Divider.UDT";
   END_VAR
BEGIN
   #divider.background_animate := "Color.String_to_DInt"("BORDER_COLOR");
   #divider.line_animate := "Color.String_to_DInt"("DIVIDER_COLOR");
END_FUNCTION

FUNCTION "Divider.Initialize" : Void   // FC46, SCL
{ S7_Optimized_Access := 'TRUE' }
VERSION : 0.1
   VAR_IN_OUT
      divider : "Divider.UDT";
   END_VAR
BEGIN
   "Divider.Show"(#divider);
   "Divider.Initialize_Colors"(#divider);
END_FUNCTION

// folder: material_hmi

FUNCTION "Material_HMI.Initialize_Display" : Void   // FC37, SCL
{ S7_Optimized_Access := 'TRUE' }
VERSION : 0.1
   VAR_IN_OUT
      material : "Materials.HMI.UDT";
   END_VAR
BEGIN
   "Screen_Background.Initialize"(#material.background);
   "Row_Data.Initialize"(#material.heat);
   "Row_Label.Initialize"(#material.header);
   "Divider.Initialize"(#material.divider);
   "Row_Data.Initialize"(#material.manganese);
   "Row_Data.Initialize"(#material.silicon);
   "Row_Data.Initialize"(#material.chromium);
   "Row_Data.Initialize"(#material.vanadium);
   "Row_Data.Initialize"(#material.nickel);
   "Row_Data.Initialize"(#material.molybdenum);
   "Row_Custom.Initialize"(#material.custom);
   "Divider.Initialize"(#material.bottom_border);
   "Divider.Hide_Line"(#material.bottom_border);
END_FUNCTION

FUNCTION "Material_HMI.Input_Animations" : Void   // FC76, SCL
{ S7_Optimized_Access := 'TRUE' }
VERSION : 0.1
   VAR_IN_OUT
      material : "Materials.HMI.UDT";
   END_VAR
BEGIN
   "Row_Data.Animate_In_Focus"(#material.heat);
   "Row_Data.Animate_In_Focus"(#material.manganese);
   "Row_Data.Animate_In_Focus"(#material.silicon);
   "Row_Data.Animate_In_Focus"(#material.chromium);
   "Row_Data.Animate_In_Focus"(#material.vanadium);
   "Row_Data.Animate_In_Focus"(#material.nickel);
   "Row_Data.Animate_In_Focus"(#material.molybdenum);
   "Row_Custom.Animate_In_Focus"(#material.custom);
END_FUNCTION

// folder: material_message

FUNCTION_BLOCK "Material_Message.Reset_Display_Driver"   // FB7, SCL
{ S7_Optimized_Access := 'TRUE' }
VERSION : 0.1
   VAR_INPUT
      send_buffer : "ADP.Message_Buffer.UDT";
   END_VAR
   VAR_IN_OUT
      interface : "Materials.HMI.UDT";
   END_VAR
   VAR
      "Message.Detect_Change_Instance" : "Message.Detect_Change";
      Reset_Display_Timer : TOF_TIME;
      old : Struct
         reset : Bool;
      END_STRUCT;
   END_VAR
   VAR_TEMP
      _message_changed : Bool;
      _et : Time;
      _reset_display : Bool;
   END_VAR
   VAR CONSTANT
      RESET_TIME : Time := T#10m;
   END_VAR
BEGIN
   #"Message.Detect_Change_Instance"(send_buffer := #send_buffer,
                                     detected := #_message_changed);
   #Reset_Display_Timer(IN := #_message_changed,
                        PT := #RESET_TIME,
                        Q => #_reset_display,
                        ET => #_et);
   IF NOT #_reset_display AND #old.reset THEN
       "Material_Message.Reset_Display"(#interface);
   END_IF;
   #old.reset := #_reset_display;
END_FUNCTION_BLOCK
